(* Logix 5000 project; controller UOWHF Emulate 5570 rev 30.12; software revision 30.00; part 9 of 13 *)
(* tags used below, declared in another part *)
   UOWHF_Add_c : DINT;
   UOWHF_Msg : DINT[16];
   UOWHF_Result : DINT[16];
(* MainProgram, continued *)

   		UOWHF_Add_c.5:=UOWHF_Result[5].31;
   		UOWHF_Result[5].31:=0;
   		UOWHF_Result[6]:=UOWHF_Result[6] + 1533867680+UOWHF_Add_c;
   		UOWHF_Add_c.6:=UOWHF_Result[6].31;
   		UOWHF_Result[6].31:=0;
   		UOWHF_Result[7]:=UOWHF_Result[7] + 1271222752+UOWHF_Add_c;
   		UOWHF_Add_c.7:=UOWHF_Result[7].31;
   		UOWHF_Result[7].31:=0;
   		UOWHF_Result[8]:=UOWHF_Result[8] + 596060815+UOWHF_Add_c;
   		UOWHF_Add_c.8:=UOWHF_Result[8].31;
   		UOWHF_Result[8].31:=0;
   	End_If;
   	If UOWHF_Msg[5].[2] Then
   		UOWHF_Result[0]:=UOWHF_Result[0] + 242207897+UOWHF_Add_c;
   		UOWHF_Add_c.0:=UOWHF_Result[0].31;
   		UOWHF_Result[0].31:=0;
   		UOWHF_Result[1]:=UOWHF_Result[1] + 1213899729+UOWHF_Add_c;
   		UOWHF_Add_c.1:=UOWHF_Result[1].31;
   		UOWHF_Result[1].31:=0;
   		UOWHF_Result[2]:=UOWHF_Result[2] + 1507311732+UOWHF_Add_c;
   		UOWHF_Add_c.2:=UOWHF_Result[2].31;
   		UOWHF_Result[2].31:=0;
   		UOWHF_Result[3]:=UOWHF_Result[3] + 850718783+UOWHF_Add_c;
   		UOWHF_Add_c.3:=UOWHF_Result[3].31;
   		UOWHF_Result[3].31:=0;
   		UOWHF_Result[4]:=UOWHF_Result[4] + 1225139163+UOWHF_Add_c;
   		UOWHF_Add_c.4:=UOWHF_Result[4].31;
   		UOWHF_Result[4].31:=0;
   		UOWHF_Result[5]:=UOWHF_Result[5] + 1524287717+UOWHF_Add_c;
   		UOWHF_Add_c.5:=UOWHF_Result[5].31;
   		UOWHF_Result[5].31:=0;
   		UOWHF_Result[6]:=UOWHF_Result[6] + 1895354303+UOWHF_Add_c;
   		UOWHF_Add_c.6:=UOWHF_Result[6].31;
   		UOWHF_Result[6].31:=0;
   		UOWHF_Result[7]:=UOWHF_Result[7] + 101628531+UOWHF_Add_c;
   		UOWHF_Add_c.7:=UOWHF_Result[7].31;
   		UOWHF_Result[7].31:=0;
   		UOWHF_Result[8]:=UOWHF_Result[8] + 114576046+UOWHF_Add_c;
   		UOWHF_Add_c.8:=UOWHF_Result[8].31;
   		UOWHF_Result[8].31:=0;
   	End_If;
   	If UOWHF_Msg[5].[3] Then
   		UOWHF_Result[0]:=UOWHF_Result[0] + 768654565+UOWHF_Add_c;
   		UOWHF_Add_c.0:=UOWHF_Result[0].31;
   		UOWHF_Result[0].31:=0;
   		UOWHF_Result[1]:=UOWHF_Result[1] + 754430999+UOWHF_Add_c;
   		UOWHF_Add_c.1:=UOWHF_Result[1].31;
   		UOWHF_Result[1].31:=0;
   		UOWHF_Result[2]:=UOWHF_Result[2] + 1940032004+UOWHF_Add_c;
   		UOWHF_Add_c.2:=UOWHF_Result[2].31;
   		UOWHF_Result[2].31:=0;
   		UOWHF_Result[3]:=UOWHF_Result[3] + 595150839+UOWHF_Add_c;
   		UOWHF_Add_c.3:=UOWHF_Result[3].31;
   		UOWHF_Result[3].31:=0;
   		UOWHF_Result[4]:=UOWHF_Result[4] + 151811053+UOWHF_Add_c;
   		UOWHF_Add_c.4:=UOWHF_Result[4].31;
   		UOWHF_Result[4].31:=0;
   		UOWHF_Result[5]:=UOWHF_Result[5] + 1466273385+UOWHF_Add_c;
   		UOWHF_Add_c.5:=UOWHF_Result[5].31;
   		UOWHF_Result[5].31:=0;
   		UOWHF_Result[6]:=UOWHF_Result[6] + 252929464+UOWHF_Add_c;
   		UOWHF_Add_c.6:=UOWHF_Result[6].31;
   		UOWHF_Result[6].31:=0;
   		UOWHF_Result[7]:=UOWHF_Result[7] + 613047462+UOWHF_Add_c;
   		UOWHF_Add_c.7:=UOWHF_Result[7].31;
   		UOWHF_Result[7].31:=0;
   		UOWHF_Result[8]:=UOWHF_Result[8] + 1252399508+UOWHF_Add_c;
   		UOWHF_Add_c.8:=UOWHF_Result[8].31;
   		UOWHF_Result[8].31:=0;
   	End_If;
   	If UOWHF_Msg[5].[4] Then
   		UOWHF_Result[0]:=UOWHF_Result[0] + 1600450797+UOWHF_Add_c;
   		UOWHF_Add_c.0:=UOWHF_Result[0].31;
   		UOWHF_Result[0].31:=0;
   		UOWHF_Result[1]:=UOWHF_Result[1] + 397376901+UOWHF_Add_c;
   		UOWHF_Add_c.1:=UOWHF_Result[1].31;
   		UOWHF_Result[1].31:=0;
   		UOWHF_Result[2]:=UOWHF_Result[2] + 844948019+UOWHF_Add_c;
   		UOWHF_Add_c.2:=UOWHF_Result[2].31;
   		UOWHF_Result[2].31:=0;
   		UOWHF_Result[3]:=UOWHF_Result[3] + 386657454+UOWHF_Add_c;
   		UOWHF_Add_c.3:=UOWHF_Result[3].31;
   		UOWHF_Result[3].31:=0;
   		UOWHF_Result[4]:=UOWHF_Result[4] + 1471910063+UOWHF_Add_c;
   		UOWHF_Add_c.4:=UOWHF_Result[4].31;
   		UOWHF_Result[4].31:=0;
   		UOWHF_Result[5]:=UOWHF_Result[5] + 162797883+UOWHF_Add_c;
   		UOWHF_Add_c.5:=UOWHF_Result[5].31;
   		UOWHF_Result[5].31:=0;
   		UOWHF_Result[6]:=UOWHF_Result[6] + 784996524+UOWHF_Add_c;
   		UOWHF_Add_c.6:=UOWHF_Result[6].31;
   		UOWHF_Result[6].31:=0;
   		UOWHF_Result[7]:=UOWHF_Result[7] + 2013933554+UOWHF_Add_c;
   		UOWHF_Add_c.7:=UOWHF_Result[7].31;
   		UOWHF_Result[7].31:=0;
   		UOWHF_Result[8]:=UOWHF_Result[8] + 440569606+UOWHF_Add_c;
   		UOWHF_Add_c.8:=UOWHF_Result[8].31;
   		UOWHF_Result[8].31:=0;
   	End_If;
   	If UOWHF_Msg[5].[5] Then
   		UOWHF_Result[0]:=UOWHF_Result[0] + 1951413431+UOWHF_Add_c;
   		UOWHF_Add_c.0:=UOWHF_Result[0].31;
   		UOWHF_Result[0].31:=0;
   		UOWHF_Result[1]:=UOWHF_Result[1] + 1309639671+UOWHF_Add_c;
   		UOWHF_Add_c.1:=UOWHF_Result[1].31;
   		UOWHF_Result[1].31:=0;
   		UOWHF_Result[2]:=UOWHF_Result[2] + 1329635265+UOWHF_Add_c;
   		UOWHF_Add_c.2:=UOWHF_Result[2].31;
   		UOWHF_Result[2].31:=0;
   		UOWHF_Result[3]:=UOWHF_Result[3] + 807074057+UOWHF_Add_c;
   		UOWHF_Add_c.3:=UOWHF_Result[3].31;
   		UOWHF_Result[3].31:=0;
   		UOWHF_Result[4]:=UOWHF_Result[4] + 1918784437+UOWHF_Add_c;
   		UOWHF_Add_c.4:=UOWHF_Result[4].31;
   		UOWHF_Result[4].31:=0;
   		UOWHF_Result[5]:=UOWHF_Result[5] + 2062494469+UOWHF_Add_c;
   		UOWHF_Add_c.5:=UOWHF_Result[5].31;
   		UOWHF_Result[5].31:=0;
   		UOWHF_Result[6]:=UOWHF_Result[6] + 472625414+UOWHF_Add_c;
   		UOWHF_Add_c.6:=UOWHF_Result[6].31;
   		UOWHF_Result[6].31:=0;
   		UOWHF_Result[7]:=UOWHF_Result[7] + 30522676+UOWHF_Add_c;
   		UOWHF_Add_c.7:=UOWHF_Result[7].31;
   		UOWHF_Result[7].31:=0;
   		UOWHF_Result[8]:=UOWHF_Result[8] + 1520794738+UOWHF_Add_c;
   		UOWHF_Add_c.8:=UOWHF_Result[8].31;
   		UOWHF_Result[8].31:=0;
   	End_If;
   	If UOWHF_Msg[5].[6] Then
   		UOWHF_Result[0]:=UOWHF_Result[0] + 627398656+UOWHF_Add_c;
   		UOWHF_Add_c.0:=UOWHF_Result[0].31;
   		UOWHF_Result[0].31:=0;
   		UOWHF_Result[1]:=UOWHF_Result[1] + 944966830+UOWHF_Add_c;
   		UOWHF_Add_c.1:=UOWHF_Result[1].31;
   		UOWHF_Result[1].31:=0;
   		UOWHF_Result[2]:=UOWHF_Result[2] + 1025387377+UOWHF_Add_c;
   		UOWHF_Add_c.2:=UOWHF_Result[2].31;
   		UOWHF_Result[2].31:=0;
   		UOWHF_Result[3]:=UOWHF_Result[3] + 713005065+UOWHF_Add_c;
   		UOWHF_Add_c.3:=UOWHF_Result[3].31;
   		UOWHF_Result[3].31:=0;
   		UOWHF_Result[4]:=UOWHF_Result[4] + 1080196444+UOWHF_Add_c;
   		UOWHF_Add_c.4:=UOWHF_Result[4].31;
   		UOWHF_Result[4].31:=0;
   		UOWHF_Result[5]:=UOWHF_Result[5] + 952605245+UOWHF_Add_c;
   		UOWHF_Add_c.5:=UOWHF_Result[5].31;
   		UOWHF_Result[5].31:=0;
   		UOWHF_Result[6]:=UOWHF_Result[6] + 1233406562+UOWHF_Add_c;
   		UOWHF_Add_c.6:=UOWHF_Result[6].31;
   		UOWHF_Result[6].31:=0;
   		UOWHF_Result[7]:=UOWHF_Result[7] + 222757426+UOWHF_Add_c;
   		UOWHF_Add_c.7:=UOWHF_Result[7].31;
   		UOWHF_Result[7].31:=0;
   		UOWHF_Result[8]:=UOWHF_Result[8] + 157633194+UOWHF_Add_c;
   		UOWHF_Add_c.8:=UOWHF_Result[8].31;
   		UOWHF_Result[8].31:=0;
   	End_If;
   	If UOWHF_Msg[5].[7] Then
   		UOWHF_Result[0]:=UOWHF_Result[0] + 1626487869+UOWHF_Add_c;
   		UOWHF_Add_c.0:=UOWHF_Result[0].31;
   		UOWHF_Result[0].31:=0;
   		UOWHF_Result[1]:=UOWHF_Result[1] + 1009587303+UOWHF_Add_c;
   		UOWHF_Add_c.1:=UOWHF_Result[1].31;
   		UOWHF_Result[1].31:=0;
   		UOWHF_Result[2]:=UOWHF_Result[2] + 2051873705+UOWHF_Add_c;
   		UOWHF_Add_c.2:=UOWHF_Result[2].31;
   		UOWHF_Result[2].31:=0;
   		UOWHF_Result[3]:=UOWHF_Result[3] + 1661358697+UOWHF_Add_c;
   		UOWHF_Add_c.3:=UOWHF_Result[3].31;
   		UOWHF_Result[3].31:=0;
   		UOWHF_Result[4]:=UOWHF_Result[4] + 275538472+UOWHF_Add_c;
   		UOWHF_Add_c.4:=UOWHF_Result[4].31;
   		UOWHF_Result[4].31:=0;
   		UOWHF_Result[5]:=UOWHF_Result[5] + 112131931+UOWHF_Add_c;
   		UOWHF_Add_c.5:=UOWHF_Result[5].31;
   		UOWHF_Result[5].31:=0;
   		UOWHF_Result[6]:=UOWHF_Result[6] + 57692083+UOWHF_Add_c;
   		UOWHF_Add_c.6:=UOWHF_Result[6].31;
   		UOWHF_Result[6].31:=0;
   		UOWHF_Result[7]:=UOWHF_Result[7] + 1369128253+UOWHF_Add_c;
   		UOWHF_Add_c.7:=UOWHF_Result[7].31;
   		UOWHF_Result[7].31:=0;
   		UOWHF_Result[8]:=UOWHF_Result[8] + 1034889855+UOWHF_Add_c;
   		UOWHF_Add_c.8:=UOWHF_Result[8].31;
   		UOWHF_Result[8].31:=0;
   	End_If;
   	If UOWHF_Msg[5].[8] Then
   		UOWHF_Result[0]:=UOWHF_Result[0] + 976942412+UOWHF_Add_c;
   		UOWHF_Add_c.0:=UOWHF_Result[0].31;
   		UOWHF_Result[0].31:=0;
   		UOWHF_Result[1]:=UOWHF_Result[1] + 711434092+UOWHF_Add_c;
   		UOWHF_Add_c.1:=UOWHF_Result[1].31;
   		UOWHF_Result[1].31:=0;
   		UOWHF_Result[2]:=UOWHF_Result[2] + 1947635793+UOWHF_Add_c;
   		UOWHF_Add_c.2:=UOWHF_Result[2].31;
   		UOWHF_Result[2].31:=0;
   		UOWHF_Result[3]:=UOWHF_Result[3] + 491121245+UOWHF_Add_c;
   		UOWHF_Add_c.3:=UOWHF_Result[3].31;
   		UOWHF_Result[3].31:=0;
   		UOWHF_Result[4]:=UOWHF_Result[4] + 1445396901+UOWHF_Add_c;
   		UOWHF_Add_c.4:=UOWHF_Result[4].31;
   		UOWHF_Result[4].31:=0;
   		UOWHF_Result[5]:=UOWHF_Result[5] + 2044325486+UOWHF_Add_c;
   		UOWHF_Add_c.5:=UOWHF_Result[5].31;
   		UOWHF_Result[5].31:=0;
   		UOWHF_Result[6]:=UOWHF_Result[6] + 1490879409+UOWHF_Add_c;
   		UOWHF_Add_c.6:=UOWHF_Result[6].31;
   		UOWHF_Result[6].31:=0;
   		UOWHF_Result[7]:=UOWHF_Result[7] + 2112785526+UOWHF_Add_c;
   		UOWHF_Add_c.7:=UOWHF_Result[7].31;
   		UOWHF_Result[7].31:=0;
   		UOWHF_Result[8]:=UOWHF_Result[8] + 392128750+UOWHF_Add_c;
   		UOWHF_Add_c.8:=UOWHF_Result[8].31;
   		UOWHF_Result[8].31:=0;
   	End_If;
   	If UOWHF_Msg[5].[9] Then
   		UOWHF_Result[0]:=UOWHF_Result[0] + 2060995341+UOWHF_Add_c;
   		UOWHF_Add_c.0:=UOWHF_Result[0].31;
   		UOWHF_Result[0].31:=0;
   		UOWHF_Result[1]:=UOWHF_Result[1] + 1687585711+UOWHF_Add_c;
   		UOWHF_Add_c.1:=UOWHF_Result[1].31;
   		UOWHF_Result[1].31:=0;
   		UOWHF_Result[2]:=UOWHF_Result[2] + 466383186+UOWHF_Add_c;
   		UOWHF_Add_c.2:=UOWHF_Result[2].31;
   		UOWHF_Result[2].31:=0;
   		UOWHF_Result[3]:=UOWHF_Result[3] + 1090651315+UOWHF_Add_c;
   		UOWHF_Add_c.3:=UOWHF_Result[3].31;
   		UOWHF_Result[3].31:=0;
   		UOWHF_Result[4]:=UOWHF_Result[4] + 533848303+UOWHF_Add_c;
   		UOWHF_Add_c.4:=UOWHF_Result[4].31;
   		UOWHF_Result[4].31:=0;
   		UOWHF_Result[5]:=UOWHF_Result[5] + 1054332536+UOWHF_Add_c;
   		UOWHF_Add_c.5:=UOWHF_Result[5].31;
   		UOWHF_Result[5].31:=0;
   		UOWHF_Result[6]:=UOWHF_Result[6] + 1013508397+UOWHF_Add_c;
   		UOWHF_Add_c.6:=UOWHF_Result[6].31;
   		UOWHF_Result[6].31:=0;
   		UOWHF_Result[7]:=UOWHF_Result[7] + 294639724+UOWHF_Add_c;
   		UOWHF_Add_c.7:=UOWHF_Result[7].31;
   		UOWHF_Result[7].31:=0;
   		UOWHF_Result[8]:=UOWHF_Result[8] + 1773956324+UOWHF_Add_c;
   		UOWHF_Add_c.8:=UOWHF_Result[8].31;
   		UOWHF_Result[8].31:=0;
   	End_If;
   	If UOWHF_Msg[5].[10] Then
   		UOWHF_Result[0]:=UOWHF_Result[0] + 1584897761+UOWHF_Add_c;
   		UOWHF_Add_c.0:=UOWHF_Result[0].31;
   		UOWHF_Result[0].31:=0;
   		UOWHF_Result[1]:=UOWHF_Result[1] + 1035971083+UOWHF_Add_c;
   		UOWHF_Add_c.1:=UOWHF_Result[1].31;
   		UOWHF_Result[1].31:=0;
   		UOWHF_Result[2]:=UOWHF_Result[2] + 663528773+UOWHF_Add_c;
   		UOWHF_Add_c.2:=UOWHF_Result[2].31;
   		UOWHF_Result[2].31:=0;
   		UOWHF_Result[3]:=UOWHF_Result[3] + 1884139568+UOWHF_Add_c;
   		UOWHF_Add_c.3:=UOWHF_Result[3].31;
   		UOWHF_Result[3].31:=0;
   		UOWHF_Result[4]:=UOWHF_Result[4] + 962334446+UOWHF_Add_c;
   		UOWHF_Add_c.4:=UOWHF_Result[4].31;
   		UOWHF_Result[4].31:=0;
   		UOWHF_Result[5]:=UOWHF_Result[5] + 909266750+UOWHF_Add_c;
   		UOWHF_Add_c.5:=UOWHF_Result[5].31;
   		UOWHF_Result[5].31:=0;
   		UOWHF_Result[6]:=UOWHF_Result[6] + 2064748270+UOWHF_Add_c;
   		UOWHF_Add_c.6:=UOWHF_Result[6].31;
   		UOWHF_Result[6].31:=0;
   		UOWHF_Result[7]:=UOWHF_Result[7] + 720877779+UOWHF_Add_c;
   		UOWHF_Add_c.7:=UOWHF_Result[7].31;
   		UOWHF_Result[7].31:=0;
   		UOWHF_Result[8]:=UOWHF_Result[8] + 1298627519+UOWHF_Add_c;
   		UOWHF_Add_c.8:=UOWHF_Result[8].31;
   		UOWHF_Result[8].31:=0;
   	End_If;
   	If UOWHF_Msg[5].[11] Then
   		UOWHF_Result[0]:=UOWHF_Result[0] + 838057991+UOWHF_Add_c;
   		UOWHF_Add_c.0:=UOWHF_Result[0].31;
   		UOWHF_Result[0].31:=0;
   		UOWHF_Result[1]:=UOWHF_Result[1] + 999112796+UOWHF_Add_c;
   		UOWHF_Add_c.1:=UOWHF_Result[1].31;
   		UOWHF_Result[1].31:=0;
   		UOWHF_Result[2]:=UOWHF_Result[2] + 514950667+UOWHF_Add_c;
   		UOWHF_Add_c.2:=UOWHF_Result[2].31;
   		UOWHF_Result[2].31:=0;
   		UOWHF_Result[3]:=UOWHF_Result[3] + 2131611961+UOWHF_Add_c;
   		UOWHF_Add_c.3:=UOWHF_Result[3].31;
   		UOWHF_Result[3].31:=0;
   		UOWHF_Result[4]:=UOWHF_Result[4] + 1984549024+UOWHF_Add_c;
   		UOWHF_Add_c.4:=UOWHF_Result[4].31;
   		UOWHF_Result[4].31:=0;
   		UOWHF_Result[5]:=UOWHF_Result[5] + 979935397+UOWHF_Add_c;
   		UOWHF_Add_c.5:=UOWHF_Result[5].31;
   		UOWHF_Result[5].31:=0;
   		UOWHF_Result[6]:=UOWHF_Result[6] + 752211313+UOWHF_Add_c;
   		UOWHF_Add_c.6:=UOWHF_Result[6].31;
   		UOWHF_Result[6].31:=0;
   		UOWHF_Result[7]:=UOWHF_Result[7] + 62917348+UOWHF_Add_c;
   		UOWHF_Add_c.7:=UOWHF_Result[7].31;
   		UOWHF_Result[7].31:=0;
   		UOWHF_Result[8]:=UOWHF_Result[8] + 1232896139+UOWHF_Add_c;
   		UOWHF_Add_c.8:=UOWHF_Result[8].31;
   		UOWHF_Result[8].31:=0;
   	End_If;
   	If UOWHF_Msg[5].[12] Then
   		UOWHF_Result[0]:=UOWHF_Result[0] + 933997728+UOWHF_Add_c;
   		UOWHF_Add_c.0:=UOWHF_Result[0].31;
   		UOWHF_Result[0].31:=0;
   		UOWHF_Result[1]:=UOWHF_Result[1] + 1740343240+UOWHF_Add_c;
   		UOWHF_Add_c.1:=UOWHF_Result[1].31;
   		UOWHF_Result[1].31:=0;
   		UOWHF_Result[2]:=UOWHF_Result[2] + 673819123+UOWHF_Add_c;
   		UOWHF_Add_c.2:=UOWHF_Result[2].31;
   		UOWHF_Result[2].31:=0;
   		UOWHF_Result[3]:=UOWHF_Result[3] + 150571982+UOWHF_Add_c;
   		UOWHF_Add_c.3:=UOWHF_Result[3].31;
   		UOWHF_Result[3].31:=0;
   		UOWHF_Result[4]:=UOWHF_Result[4] + 1634031125+UOWHF_Add_c;
   		UOWHF_Add_c.4:=UOWHF_Result[4].31;
   		UOWHF_Result[4].31:=0;
   		UOWHF_Result[5]:=UOWHF_Result[5] + 889194862+UOWHF_Add_c;
   		UOWHF_Add_c.5:=UOWHF_Result[5].31;
   		UOWHF_Result[5].31:=0;
   		UOWHF_Result[6]:=UOWHF_Result[6] + 1077160835+UOWHF_Add_c;
   		UOWHF_Add_c.6:=UOWHF_Result[6].31;
   		UOWHF_Result[6].31:=0;
   		UOWHF_Result[7]:=UOWHF_Result[7] + 648021849+UOWHF_Add_c;
   		UOWHF_Add_c.7:=UOWHF_Result[7].31;
   		UOWHF_Result[7].31:=0;
   		UOWHF_Result[8]:=UOWHF_Result[8] + 499612356+UOWHF_Add_c;
   		UOWHF_Add_c.8:=UOWHF_Result[8].31;
   		UOWHF_Result[8].31:=0;
   	End_If;
   	If UOWHF_Msg[5].[13] Then
   		UOWHF_Result[0]:=UOWHF_Result[0] + 98910495+UOWHF_Add_c;
   		UOWHF_Add_c.0:=UOWHF_Result[0].31;
   		UOWHF_Result[0].31:=0;
   		UOWHF_Result[1]:=UOWHF_Result[1] + 1692366771+UOWHF_Add_c;
   		UOWHF_Add_c.1:=UOWHF_Result[1].31;
   		UOWHF_Result[1].31:=0;
   		UOWHF_Result[2]:=UOWHF_Result[2] + 1102242537+UOWHF_Add_c;
   		UOWHF_Add_c.2:=UOWHF_Result[2].31;
   		UOWHF_Result[2].31:=0;
   		UOWHF_Result[3]:=UOWHF_Result[3] + 976987602+UOWHF_Add_c;
   		UOWHF_Add_c.3:=UOWHF_Result[3].31;
   		UOWHF_Result[3].31:=0;
   		UOWHF_Result[4]:=UOWHF_Result[4] + 195497023+UOWHF_Add_c;
   		UOWHF_Add_c.4:=UOWHF_Result[4].31;
   		UOWHF_Result[4].31:=0;
   		UOWHF_Result[5]:=UOWHF_Result[5] + 1969565650+UOWHF_Add_c;
   		UOWHF_Add_c.5:=UOWHF_Result[5].31;
   		UOWHF_Result[5].31:=0;
   		UOWHF_Result[6]:=UOWHF_Result[6] + 916579574+UOWHF_Add_c;
   		UOWHF_Add_c.6:=UOWHF_Result[6].31;
   		UOWHF_Result[6].31:=0;
   		UOWHF_Result[7]:=UOWHF_Result[7] + 1976862514+UOWHF_Add_c;
   		UOWHF_Add_c.7:=UOWHF_Result[7].31;
   		UOWHF_Result[7].31:=0;
   		UOWHF_Result[8]:=UOWHF_Result[8] + 251699664+UOWHF_Add_c;
   		UOWHF_Add_c.8:=UOWHF_Result[8].31;
   		UOWHF_Result[8].31:=0;
   	End_If;
   	If UOWHF_Msg[5].[14] Then
   		UOWHF_Result[0]:=UOWHF_Result[0] + 1883670867+UOWHF_Add_c;
   		UOWHF_Add_c.0:=UOWHF_Result[0].31;
   		UOWHF_Result[0].31:=0;
   		UOWHF_Result[1]:=UOWHF_Result[1] + 881302118+UOWHF_Add_c;
   		UOWHF_Add_c.1:=UOWHF_Result[1].31;
   		UOWHF_Result[1].31:=0;
   		UOWHF_Result[2]:=UOWHF_Result[2] + 646224306+UOWHF_Add_c;
   		UOWHF_Add_c.2:=UOWHF_Result[2].31;
   		UOWHF_Result[2].31:=0;
   		UOWHF_Result[3]:=UOWHF_Result[3] + 182806481+UOWHF_Add_c;
   		UOWHF_Add_c.3:=UOWHF_Result[3].31;
   		UOWHF_Result[3].31:=0;
   		UOWHF_Result[4]:=UOWHF_Result[4] + 1574869751+UOWHF_Add_c;
   		UOWHF_Add_c.4:=UOWHF_Result[4].31;
   		UOWHF_Result[4].31:=0;
   		UOWHF_Result[5]:=UOWHF_Result[5] + 216878236+UOWHF_Add_c;
   		UOWHF_Add_c.5:=UOWHF_Result[5].31;
   		UOWHF_Result[5].31:=0;
   		UOWHF_Result[6]:=UOWHF_Result[6] + 1309703789+UOWHF_Add_c;
   		UOWHF_Add_c.6:=UOWHF_Result[6].31;
   		UOWHF_Result[6].31:=0;
   		UOWHF_Result[7]:=UOWHF_Result[7] + 10544512+UOWHF_Add_c;
   		UOWHF_Add_c.7:=UOWHF_Result[7].31;
   		UOWHF_Result[7].31:=0;
   		UOWHF_Result[8]:=UOWHF_Result[8] + 1438861351+UOWHF_Add_c;
   		UOWHF_Add_c.8:=UOWHF_Result[8].31;
   		UOWHF_Result[8].31:=0;
   	End_If;
   	If UOWHF_Msg[5].[15] Then
   		UOWHF_Result[0]:=UOWHF_Result[0] + 1175849528+UOWHF_Add_c;
   		UOWHF_Add_c.0:=UOWHF_Result[0].31;
   		UOWHF_Result[0].31:=0;
   		UOWHF_Result[1]:=UOWHF_Result[1] + 593969039+UOWHF_Add_c;
   		UOWHF_Add_c.1:=UOWHF_Result[1].31;
   		UOWHF_Result[1].31:=0;
   		UOWHF_Result[2]:=UOWHF_Result[2] + 1047920593+UOWHF_Add_c;
   		UOWHF_Add_c.2:=UOWHF_Result[2].31;
   		UOWHF_Result[2].31:=0;
   		UOWHF_Result[3]:=UOWHF_Result[3] + 435488860+UOWHF_Add_c;
   		UOWHF_Add_c.3:=UOWHF_Result[3].31;
   		UOWHF_Result[3].31:=0;
   		UOWHF_Result[4]:=UOWHF_Result[4] + 2047652892+UOWHF_Add_c;
   		UOWHF_Add_c.4:=UOWHF_Result[4].31;
   		UOWHF_Result[4].31:=0;
   		UOWHF_Result[5]:=UOWHF_Result[5] + 946271868+UOWHF_Add_c;
   		UOWHF_Add_c.5:=UOWHF_Result[5].31;
   		UOWHF_Result[5].31:=0;
   		UOWHF_Result[6]:=UOWHF_Result[6] + 111644338+UOWHF_Add_c;
   		UOWHF_Add_c.6:=UOWHF_Result[6].31;
   		UOWHF_Result[6].31:=0;
   		UOWHF_Result[7]:=UOWHF_Result[7] + 697600493+UOWHF_Add_c;
   		UOWHF_Add_c.7:=UOWHF_Result[7].31;
   		UOWHF_Result[7].31:=0;
   		UOWHF_Result[8]:=UOWHF_Result[8] + 521259784+UOWHF_Add_c;
   		UOWHF_Add_c.8:=UOWHF_Result[8].31;
   		UOWHF_Result[8].31:=0;
   	End_If;
   	If UOWHF_Msg[5].[16] Then
   		UOWHF_Result[0]:=UOWHF_Result[0] + 1395198064+UOWHF_Add_c;
   		UOWHF_Add_c.0:=UOWHF_Result[0].31;
   		UOWHF_Result[0].31:=0;
   		UOWHF_Result[1]:=UOWHF_Result[1] + 1066351934+UOWHF_Add_c;
   		UOWHF_Add_c.1:=UOWHF_Result[1].31;
   		UOWHF_Result[1].31:=0;
   		UOWHF_Result[2]:=UOWHF_Result[2] + 1276681201+UOWHF_Add_c;
   		UOWHF_Add_c.2:=UOWHF_Result[2].31;
   		UOWHF_Result[2].31:=0;
   		UOWHF_Result[3]:=UOWHF_Result[3] + 80726074+UOWHF_Add_c;
   		UOWHF_Add_c.3:=UOWHF_Result[3].31;
   		UOWHF_Result[3].31:=0;
   		UOWHF_Result[4]:=UOWHF_Result[4] + 896217188+UOWHF_Add_c;
   		UOWHF_Add_c.4:=UOWHF_Result[4].31;
   		UOWHF_Result[4].31:=0;
   		UOWHF_Result[5]:=UOWHF_Result[5] + 38350786+UOWHF_Add_c;
   		UOWHF_Add_c.5:=UOWHF_Result[5].31;
   		UOWHF_Result[5].31:=0;
   		UOWHF_Result[6]:=UOWHF_Result[6] + 575258542+UOWHF_Add_c;
   		UOWHF_Add_c.6:=UOWHF_Result[6].31;
   		UOWHF_Result[6].31:=0;
   		UOWHF_Result[7]:=UOWHF_Result[7] + 499314129+UOWHF_Add_c;
   		UOWHF_Add_c.7:=UOWHF_Result[7].31;
   		UOWHF_Result[7].31:=0;
   		UOWHF_Result[8]:=UOWHF_Result[8] + 736790724+UOWHF_Add_c;
   		UOWHF_Add_c.8:=UOWHF_Result[8].31;
   		UOWHF_Result[8].31:=0;
   	End_If;
   	If UOWHF_Msg[5].[17] Then
   		UOWHF_Result[0]:=UOWHF_Result[0] + 309344076+UOWHF_Add_c;
   		UOWHF_Add_c.0:=UOWHF_Result[0].31;
   		UOWHF_Result[0].31:=0;
   		UOWHF_Result[1]:=UOWHF_Result[1] + 799987601+UOWHF_Add_c;
   		UOWHF_Add_c.1:=UOWHF_Result[1].31;
   		UOWHF_Result[1].31:=0;
   		UOWHF_Result[2]:=UOWHF_Result[2] + 1787238195+UOWHF_Add_c;
   		UOWHF_Add_c.2:=UOWHF_Result[2].31;
   		UOWHF_Result[2].31:=0;
   		UOWHF_Result[3]:=UOWHF_Result[3] + 1444841006+UOWHF_Add_c;
   		UOWHF_Add_c.3:=UOWHF_Result[3].31;
   		UOWHF_Result[3].31:=0;
   		UOWHF_Result[4]:=UOWHF_Result[4] + 716956811+UOWHF_Add_c;
   		UOWHF_Add_c.4:=UOWHF_Result[4].31;
   		UOWHF_Result[4].31:=0;
   		UOWHF_Result[5]:=UOWHF_Result[5] + 2050078126+UOWHF_Add_c;
   		UOWHF_Add_c.5:=UOWHF_Result[5].31;
   		UOWHF_Result[5].31:=0;
   		UOWHF_Result[6]:=UOWHF_Result[6] + 354965748+UOWHF_Add_c;
   		UOWHF_Add_c.6:=UOWHF_Result[6].31;
   		UOWHF_Result[6].31:=0;
   		UOWHF_Result[7]:=UOWHF_Result[7] + 696362392+UOWHF_Add_c;
   		UOWHF_Add_c.7:=UOWHF_Result[7].31;
   		UOWHF_Result[7].31:=0;
   		UOWHF_Result[8]:=UOWHF_Result[8] + 826540150+UOWHF_Add_c;
   		UOWHF_Add_c.8:=UOWHF_Result[8].31;
   		UOWHF_Result[8].31:=0;
   	End_If;
   	If UOWHF_Msg[5].[18] Then
   		UOWHF_Result[0]:=UOWHF_Result[0] + 1307778602+UOWHF_Add_c;
   		UOWHF_Add_c.0:=UOWHF_Result[0].31;
   		UOWHF_Result[0].31:=0;
   		UOWHF_Result[1]:=UOWHF_Result[1] + 2143863024+UOWHF_Add_c;
   		UOWHF_Add_c.1:=UOWHF_Result[1].31;
   		UOWHF_Result[1].31:=0;
   		UOWHF_Result[2]:=UOWHF_Result[2] + 1414502428+UOWHF_Add_c;
   		UOWHF_Add_c.2:=UOWHF_Result[2].31;
   		UOWHF_Result[2].31:=0;
   		UOWHF_Result[3]:=UOWHF_Result[3] + 555690590+UOWHF_Add_c;
   		UOWHF_Add_c.3:=UOWHF_Result[3].31;
   		UOWHF_Result[3].31:=0;
   		UOWHF_Result[4]:=UOWHF_Result[4] + 149275133+UOWHF_Add_c;
   		UOWHF_Add_c.4:=UOWHF_Result[4].31;
   		UOWHF_Result[4].31:=0;
   		UOWHF_Result[5]:=UOWHF_Result[5] + 914353412+UOWHF_Add_c;
   		UOWHF_Add_c.5:=UOWHF_Result[5].31;
   		UOWHF_Result[5].31:=0;
   		UOWHF_Result[6]:=UOWHF_Result[6] + 1687495362+UOWHF_Add_c;
   		UOWHF_Add_c.6:=UOWHF_Result[6].31;
   		UOWHF_Result[6].31:=0;
   		UOWHF_Result[7]:=UOWHF_Result[7] + 104151502+UOWHF_Add_c;
   		UOWHF_Add_c.7:=UOWHF_Result[7].31;
   		UOWHF_Result[7].31:=0;
   		UOWHF_Result[8]:=UOWHF_Result[8] + 1701136503+UOWHF_Add_c;
   		UOWHF_Add_c.8:=UOWHF_Result[8].31;
   		UOWHF_Result[8].31:=0;
   	End_If;
   	If UOWHF_Msg[5].[19] Then
   		UOWHF_Result[0]:=UOWHF_Result[0] + 728052003+UOWHF_Add_c;
   		UOWHF_Add_c.0:=UOWHF_Result[0].31;
   		UOWHF_Result[0].31:=0;
   		UOWHF_Result[1]:=UOWHF_Result[1] + 2107753207+UOWHF_Add_c;
   		UOWHF_Add_c.1:=UOWHF_Result[1].31;
   		UOWHF_Result[1].31:=0;
   		UOWHF_Result[2]:=UOWHF_Result[2] + 971727159+UOWHF_Add_c;
   		UOWHF_Add_c.2:=UOWHF_Result[2].31;
   		UOWHF_Result[2].31:=0;
   		UOWHF_Result[3]:=UOWHF_Result[3] + 1190530007+UOWHF_Add_c;
   		UOWHF_Add_c.3:=UOWHF_Result[3].31;
   		UOWHF_Result[3].31:=0;
   		UOWHF_Result[4]:=UOWHF_Result[4] + 1927683191+UOWHF_Add_c;
   		UOWHF_Add_c.4:=UOWHF_Result[4].31;
   		UOWHF_Result[4].31:=0;
   		UOWHF_Result[5]:=UOWHF_Result[5] + 1162645362+UOWHF_Add_c;
   		UOWHF_Add_c.5:=UOWHF_Result[5].31;
   		UOWHF_Result[5].31:=0;
   		UOWHF_Result[6]:=UOWHF_Result[6] + 2123028397+UOWHF_Add_c;
   		UOWHF_Add_c.6:=UOWHF_Result[6].31;
   		UOWHF_Result[6].31:=0;
   		UOWHF_Result[7]:=UOWHF_Result[7] + 1950322746+UOWHF_Add_c;
   		UOWHF_Add_c.7:=UOWHF_Result[7].31;
   		UOWHF_Result[7].31:=0;
   		UOWHF_Result[8]:=UOWHF_Result[8] + 468197333+UOWHF_Add_c;
   		UOWHF_Add_c.8:=UOWHF_Result[8].31;
   		UOWHF_Result[8].31:=0;
   	End_If;
   	If UOWHF_Msg[5].[20] Then
   		UOWHF_Result[0]:=UOWHF_Result[0] + 92482565+UOWHF_Add_c;
   		UOWHF_Add_c.0:=UOWHF_Result[0].31;
   		UOWHF_Result[0].31:=0;
   		UOWHF_Result[1]:=UOWHF_Result[1] + 659136073+UOWHF_Add_c;
   		UOWHF_Add_c.1:=UOWHF_Result[1].31;
   		UOWHF_Result[1].31:=0;
   		UOWHF_Result[2]:=UOWHF_Result[2] + 1245607757+UOWHF_Add_c;
   		UOWHF_Add_c.2:=UOWHF_Result[2].31;
   		UOWHF_Result[2].31:=0;
   		UOWHF_Result[3]:=UOWHF_Result[3] + 1663935487+UOWHF_Add_c;
   		UOWHF_Add_c.3:=UOWHF_Result[3].31;
   		UOWHF_Result[3].31:=0;
   		UOWHF_Result[4]:=UOWHF_Result[4] + 585571943+UOWHF_Add_c;
   		UOWHF_Add_c.4:=UOWHF_Result[4].31;
   		UOWHF_Result[4].31:=0;
   		UOWHF_Result[5]:=UOWHF_Result[5] + 88073602+UOWHF_Add_c;
   		UOWHF_Add_c.5:=UOWHF_Result[5].31;
   		UOWHF_Result[5].31:=0;
   		UOWHF_Result[6]:=UOWHF_Result[6] + 2043878638+UOWHF_Add_c;
   		UOWHF_Add_c.6:=UOWHF_Result[6].31;
   		UOWHF_Result[6].31:=0;
   		UOWHF_Result[7]:=UOWHF_Result[7] + 978762805+UOWHF_Add_c;
   		UOWHF_Add_c.7:=UOWHF_Result[7].31;
   		UOWHF_Result[7].31:=0;
   		UOWHF_Result[8]:=UOWHF_Result[8] + 142446245+UOWHF_Add_c;
   		UOWHF_Add_c.8:=UOWHF_Result[8].31;
   		UOWHF_Result[8].31:=0;
   	End_If;
   	If UOWHF_Msg[5].[21] Then
   		UOWHF_Result[0]:=UOWHF_Result[0] + 1326621747+UOWHF_Add_c;
   		UOWHF_Add_c.0:=UOWHF_Result[0].31;
   		UOWHF_Result[0].31:=0;
   		UOWHF_Result[1]:=UOWHF_Result[1] + 1527242615+UOWHF_Add_c;
   		UOWHF_Add_c.1:=UOWHF_Result[1].31;
   		UOWHF_Result[1].31:=0;
   		UOWHF_Result[2]:=UOWHF_Result[2] + 1036610998+UOWHF_Add_c;
   		UOWHF_Add_c.2:=UOWHF_Result[2].31;
   		UOWHF_Result[2].31:=0;
   		UOWHF_Result[3]:=UOWHF_Result[3] + 2106304214+UOWHF_Add_c;
   		UOWHF_Add_c.3:=UOWHF_Result[3].31;
   		UOWHF_Result[3].31:=0;
   		UOWHF_Result[4]:=UOWHF_Result[4] + 1622504932+UOWHF_Add_c;
   		UOWHF_Add_c.4:=UOWHF_Result[4].31;
   		UOWHF_Result[4].31:=0;
   		UOWHF_Result[5]:=UOWHF_Result[5] + 950916145+UOWHF_Add_c;
   		UOWHF_Add_c.5:=UOWHF_Result[5].31;
   		UOWHF_Result[5].31:=0;
   		UOWHF_Result[6]:=UOWHF_Result[6] + 1107607354+UOWHF_Add_c;
   		UOWHF_Add_c.6:=UOWHF_Result[6].31;
   		UOWHF_Result[6].31:=0;
   		UOWHF_Result[7]:=UOWHF_Result[7] + 711119777+UOWHF_Add_c;
   		UOWHF_Add_c.7:=UOWHF_Result[7].31;
   		UOWHF_Result[7].31:=0;
   		UOWHF_Result[8]:=UOWHF_Result[8] + 563440627+UOWHF_Add_c;
   		UOWHF_Add_c.8:=UOWHF_Result[8].31;
   		UOWHF_Result[8].31:=0;
   	End_If;
   	If UOWHF_Msg[5].[22] Then
   		UOWHF_Result[0]:=UOWHF_Result[0] + 1902098681+UOWHF_Add_c;
   		UOWHF_Add_c.0:=UOWHF_Result[0].31;
   		UOWHF_Result[0].31:=0;
   		UOWHF_Result[1]:=UOWHF_Result[1] + 1896466664+UOWHF_Add_c;
   		UOWHF_Add_c.1:=UOWHF_Result[1].31;
   		UOWHF_Result[1].31:=0;
   		UOWHF_Result[2]:=UOWHF_Result[2] + 662408686+UOWHF_Add_c;
   		UOWHF_Add_c.2:=UOWHF_Result[2].31;
   		UOWHF_Result[2].31:=0;
   		UOWHF_Result[3]:=UOWHF_Result[3] + 2038779258+UOWHF_Add_c;
   		UOWHF_Add_c.3:=UOWHF_Result[3].31;
   		UOWHF_Result[3].31:=0;
   		UOWHF_Result[4]:=UOWHF_Result[4] + 2046912342+UOWHF_Add_c;
   		UOWHF_Add_c.4:=UOWHF_Result[4].31;
   		UOWHF_Result[4].31:=0;
   		UOWHF_Result[5]:=UOWHF_Result[5] + 585042939+UOWHF_Add_c;
   		UOWHF_Add_c.5:=UOWHF_Result[5].31;
   		UOWHF_Result[5].31:=0;
   		UOWHF_Result[6]:=UOWHF_Result[6] + 533830927+UOWHF_Add_c;
   		UOWHF_Add_c.6:=UOWHF_Result[6].31;
   		UOWHF_Result[6].31:=0;
   		UOWHF_Result[7]:=UOWHF_Result[7] + 1835939803+UOWHF_Add_c;
   		UOWHF_Add_c.7:=UOWHF_Result[7].31;
   		UOWHF_Result[7].31:=0;
   		UOWHF_Result[8]:=UOWHF_Result[8] + 736661196+UOWHF_Add_c;
   		UOWHF_Add_c.8:=UOWHF_Result[8].31;
   		UOWHF_Result[8].31:=0;
   	End_If;
   	If UOWHF_Msg[5].[23] Then
   		UOWHF_Result[0]:=UOWHF_Result[0] + 1248316559+UOWHF_Add_c;
   		UOWHF_Add_c.0:=UOWHF_Result[0].31;
   		UOWHF_Result[0].31:=0;
   		UOWHF_Result[1]:=UOWHF_Result[1] + 1056227022+UOWHF_Add_c;
   		UOWHF_Add_c.1:=UOWHF_Result[1].31;
   		UOWHF_Result[1].31:=0;
   		UOWHF_Result[2]:=UOWHF_Result[2] + 6347178+UOWHF_Add_c;
   		UOWHF_Add_c.2:=UOWHF_Result[2].31;
   		UOWHF_Result[2].31:=0;
   		UOWHF_Result[3]:=UOWHF_Result[3] + 473297225+UOWHF_Add_c;
   		UOWHF_Add_c.3:=UOWHF_Result[3].31;
   		UOWHF_Result[3].31:=0;
   		UOWHF_Result[4]:=UOWHF_Result[4] + 1833441285+UOWHF_Add_c;
   		UOWHF_Add_c.4:=UOWHF_Result[4].31;
   		UOWHF_Result[4].31:=0;
   		UOWHF_Result[5]:=UOWHF_Result[5] + 1052507972+UOWHF_Add_c;
   		UOWHF_Add_c.5:=UOWHF_Result[5].31;
   		UOWHF_Result[5].31:=0;
   		UOWHF_Result[6]:=UOWHF_Result[6] + 703965614+UOWHF_Add_c;
   		UOWHF_Add_c.6:=UOWHF_Result[6].31;
   		UOWHF_Result[6].31:=0;
   		UOWHF_Result[7]:=UOWHF_Result[7] + 807679768+UOWHF_Add_c;
   		UOWHF_Add_c.7:=UOWHF_Result[7].31;
   		UOWHF_Result[7].31:=0;
   		UOWHF_Result[8]:=UOWHF_Result[8] + 1331801305+UOWHF_Add_c;
   		UOWHF_Add_c.8:=UOWHF_Result[8].31;
   		UOWHF_Result[8].31:=0;
   	End_If;
   	If UOWHF_Msg[5].[24] Then
   		UOWHF_Result[0]:=UOWHF_Result[0] + 1719074991+UOWHF_Add_c;
   		UOWHF_Add_c.0:=UOWHF_Result[0].31;
   		UOWHF_Result[0].31:=0;
   		UOWHF_Result[1]:=UOWHF_Result[1] + 1812051904+UOWHF_Add_c;
   		UOWHF_Add_c.1:=UOWHF_Result[1].31;
   		UOWHF_Result[1].31:=0;
   		UOWHF_Result[2]:=UOWHF_Result[2] + 307015602+UOWHF_Add_c;
   		UOWHF_Add_c.2:=UOWHF_Result[2].31;
   		UOWHF_Result[2].31:=0;
   		UOWHF_Result[3]:=UOWHF_Result[3] + 180972567+UOWHF_Add_c;
   		UOWHF_Add_c.3:=UOWHF_Result[3].31;
   		UOWHF_Result[3].31:=0;
   		UOWHF_Result[4]:=UOWHF_Result[4] + 1531392063+UOWHF_Add_c;
   		UOWHF_Add_c.4:=UOWHF_Result[4].31;
   		UOWHF_Result[4].31:=0;
   		UOWHF_Result[5]:=UOWHF_Result[5] + 336776407+UOWHF_Add_c;
   		UOWHF_Add_c.5:=UOWHF_Result[5].31;
   		UOWHF_Result[5].31:=0;
   		UOWHF_Result[6]:=UOWHF_Result[6] + 189360354+UOWHF_Add_c;
   		UOWHF_Add_c.6:=UOWHF_Result[6].31;
   		UOWHF_Result[6].31:=0;
   		UOWHF_Result[7]:=UOWHF_Result[7] + 821930879+UOWHF_Add_c;
   		UOWHF_Add_c.7:=UOWHF_Result[7].31;
   		UOWHF_Result[7].31:=0;
   		UOWHF_Result[8]:=UOWHF_Result[8] + 848215891+UOWHF_Add_c;
   		UOWHF_Add_c.8:=UOWHF_Result[8].31;
   		UOWHF_Result[8].31:=0;
   	End_If;
   	If UOWHF_Msg[5].[25] Then
   		UOWHF_Result[0]:=UOWHF_Result[0] + 878116638+UOWHF_Add_c;
   		UOWHF_Add_c.0:=UOWHF_Result[0].31;
   		UOWHF_Result[0].31:=0;
   		UOWHF_Result[1]:=UOWHF_Result[1] + 1696922735+UOWHF_Add_c;
   		UOWHF_Add_c.1:=UOWHF_Result[1].31;
   		UOWHF_Result[1].31:=0;
   		UOWHF_Result[2]:=UOWHF_Result[2] + 846929162+UOWHF_Add_c;
   		UOWHF_Add_c.2:=UOWHF_Result[2].31;
   		UOWHF_Result[2].31:=0;
   		UOWHF_Result[3]:=UOWHF_Result[3] + 590335165+UOWHF_Add_c;
   		UOWHF_Add_c.3:=UOWHF_Result[3].31;
   		UOWHF_Result[3].31:=0;
   		UOWHF_Result[4]:=UOWHF_Result[4] + 950264241+UOWHF_Add_c;
   		UOWHF_Add_c.4:=UOWHF_Result[4].31;
   		UOWHF_Result[4].31:=0;
   		UOWHF_Result[5]:=UOWHF_Result[5] + 1372255350+UOWHF_Add_c;
   		UOWHF_Add_c.5:=UOWHF_Result[5].31;
   		UOWHF_Result[5].31:=0;
   		UOWHF_Result[6]:=UOWHF_Result[6] + 375515807+UOWHF_Add_c;
   		UOWHF_Add_c.6:=UOWHF_Result[6].31;
   		UOWHF_Result[6].31:=0;
   		UOWHF_Result[7]:=UOWHF_Result[7] + 2071216937+UOWHF_Add_c;
   		UOWHF_Add_c.7:=UOWHF_Result[7].31;
   		UOWHF_Result[7].31:=0;
   		UOWHF_Result[8]:=UOWHF_Result[8] + 99390644+UOWHF_Add_c;
   		UOWHF_Add_c.8:=UOWHF_Result[8].31;
   		UOWHF_Result[8].31:=0;
   	End_If;
   	If UOWHF_Msg[5].[26] Then
   		UOWHF_Result[0]:=UOWHF_Result[0] + 1005669034+UOWHF_Add_c;
   		UOWHF_Add_c.0:=UOWHF_Result[0].31;
   		UOWHF_Result[0].31:=0;
   		UOWHF_Result[1]:=UOWHF_Result[1] + 1011993720+UOWHF_Add_c;
   		UOWHF_Add_c.1:=UOWHF_Result[1].31;
   		UOWHF_Result[1].31:=0;
   		UOWHF_Result[2]:=UOWHF_Result[2] + 1387484612+UOWHF_Add_c;
   		UOWHF_Add_c.2:=UOWHF_Result[2].31;
   		UOWHF_Result[2].31:=0;
   		UOWHF_Result[3]:=UOWHF_Result[3] + 510210382+UOWHF_Add_c;
   		UOWHF_Add_c.3:=UOWHF_Result[3].31;
   		UOWHF_Result[3].31:=0;
   		UOWHF_Result[4]:=UOWHF_Result[4] + 989828960+UOWHF_Add_c;
   		UOWHF_Add_c.4:=UOWHF_Result[4].31;
   		UOWHF_Result[4].31:=0;
   		UOWHF_Result[5]:=UOWHF_Result[5] + 1812403662+UOWHF_Add_c;
   		UOWHF_Add_c.5:=UOWHF_Result[5].31;
   		UOWHF_Result[5].31:=0;
   		UOWHF_Result[6]:=UOWHF_Result[6] + 2138870626+UOWHF_Add_c;
   		UOWHF_Add_c.6:=UOWHF_Result[6].31;
   		UOWHF_Result[6].31:=0;
   		UOWHF_Result[7]:=UOWHF_Result[7] + 1448647192+UOWHF_Add_c;
   		UOWHF_Add_c.7:=UOWHF_Result[7].31;
   		UOWHF_Result[7].31:=0;
   		UOWHF_Result[8]:=UOWHF_Result[8] + 1732892583+UOWHF_Add_c;
   		UOWHF_Add_c.8:=UOWHF_Result[8].31;
   		UOWHF_Result[8].31:=0;
   	End_If;
   	If UOWHF_Msg[5].[27] Then
   		UOWHF_Result[0]:=UOWHF_Result[0] + 651670476+UOWHF_Add_c;
   		UOWHF_Add_c.0:=UOWHF_Result[0].31;
   		UOWHF_Result[0].31:=0;
   		UOWHF_Result[1]:=UOWHF_Result[1] + 1354131750+UOWHF_Add_c;
   		UOWHF_Add_c.1:=UOWHF_Result[1].31;
   		UOWHF_Result[1].31:=0;
   		UOWHF_Result[2]:=UOWHF_Result[2] + 708585138+UOWHF_Add_c;
   		UOWHF_Add_c.2:=UOWHF_Result[2].31;
   		UOWHF_Result[2].31:=0;
   		UOWHF_Result[3]:=UOWHF_Result[3] + 20236604+UOWHF_Add_c;
   		UOWHF_Add_c.3:=UOWHF_Result[3].31;
   		UOWHF_Result[3].31:=0;
   		UOWHF_Result[4]:=UOWHF_Result[4] + 155160992+UOWHF_Add_c;
   		UOWHF_Add_c.4:=UOWHF_Result[4].31;
   		UOWHF_Result[4].31:=0;
   		UOWHF_Result[5]:=UOWHF_Result[5] + 1727729102+UOWHF_Add_c;
   		UOWHF_Add_c.5:=UOWHF_Result[5].31;
   		UOWHF_Result[5].31:=0;
   		UOWHF_Result[6]:=UOWHF_Result[6] + 871695250+UOWHF_Add_c;
   		UOWHF_Add_c.6:=UOWHF_Result[6].31;
   		UOWHF_Result[6].31:=0;
   		UOWHF_Result[7]:=UOWHF_Result[7] + 1011547996+UOWHF_Add_c;
   		UOWHF_Add_c.7:=UOWHF_Result[7].31;
   		UOWHF_Result[7].31:=0;
   		UOWHF_Result[8]:=UOWHF_Result[8] + 1391268742+UOWHF_Add_c;
   		UOWHF_Add_c.8:=UOWHF_Result[8].31;
   		UOWHF_Result[8].31:=0;
   	End_If;
   	If UOWHF_Msg[5].[28] Then
   		UOWHF_Result[0]:=UOWHF_Result[0] + 2048508856+UOWHF_Add_c;
   		UOWHF_Add_c.0:=UOWHF_Result[0].31;
   		UOWHF_Result[0].31:=0;
   		UOWHF_Result[1]:=UOWHF_Result[1] + 706161872+UOWHF_Add_c;
   		UOWHF_Add_c.1:=UOWHF_Result[1].31;
   		UOWHF_Result[1].31:=0;
   		UOWHF_Result[2]:=UOWHF_Result[2] + 1143431411+UOWHF_Add_c;
   		UOWHF_Add_c.2:=UOWHF_Result[2].31;
   		UOWHF_Result[2].31:=0;
   		UOWHF_Result[3]:=UOWHF_Result[3] + 902991407+UOWHF_Add_c;
   		UOWHF_Add_c.3:=UOWHF_Result[3].31;